// TIA Portal project "FORMING_1500_PLC" (V15) (continued)

REGION Network 7: Q124.4 ON SELAMA 6 DETIK SETELAH I 7.5 ON
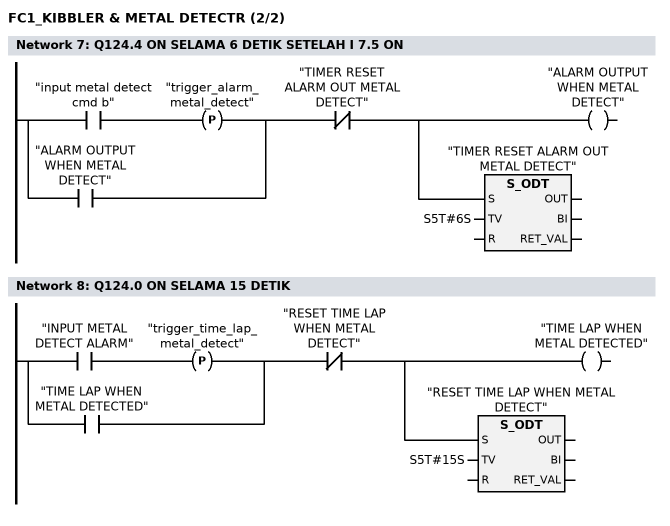
   RUNG wire#powerrail
      Contact( "input metal detect cmd b" )
      P_Trig( "trigger_alarm_metal_detect" )
      wire#w1
      I_Contact( "TIMER RESET ALARM OUT METAL DETECT" )
      wire#w2
      Coil( "ALARM OUTPUT WHEN METAL DETECT" )
   END_RUNG
   RUNG wire#powerrail
      Contact( "ALARM OUTPUT WHEN METAL DETECT" )
   END_RUNG wire#w1
   RUNG wire#w2
      S_ODT(T_NO := "TIMER RESET ALARM OUT METAL DETECT", TV := S5T#6S, R :=, BI =>, RET_VAL =>)
   END_RUNG
   // the same network as SCL:
   #_w1 := "input metal detect cmd b" AND NOT "trigger_alarm_metal_detect";   // rising edge
   "trigger_alarm_metal_detect" := "input metal detect cmd b";
   "ALARM OUTPUT WHEN METAL DETECT" := (#_w1 OR "ALARM OUTPUT WHEN METAL DETECT") AND NOT "TIMER RESET ALARM OUT METAL DETECT";
   #_s5time1 := S_ODT(T_NO := "TIMER RESET ALARM OUT METAL DETECT",
                      S := "ALARM OUTPUT WHEN METAL DETECT",
                      TV := S5T#6S);
END_REGION

REGION Network 8: Q124.0 ON SELAMA 15 DETIK
   RUNG wire#powerrail
      Contact( "INPUT METAL DETECT ALARM" )
      P_Trig( "trigger_time_lap_metal_detect" )
      wire#w1
      I_Contact( "RESET TIME LAP WHEN METAL DETECT" )
      wire#w2
      Coil( "TIME LAP WHEN METAL DETECTED" )
   END_RUNG
   RUNG wire#powerrail
      Contact( "TIME LAP WHEN METAL DETECTED" )
   END_RUNG wire#w1
   RUNG wire#w2
      S_ODT(T_NO := "RESET TIME LAP WHEN METAL DETECT", TV := S5T#15S, R :=, BI =>, RET_VAL =>)
   END_RUNG
   // the same network as SCL:
   #_w1 := "INPUT METAL DETECT ALARM" AND NOT "trigger_time_lap_metal_detect";   // rising edge
   "trigger_time_lap_metal_detect" := "INPUT METAL DETECT ALARM";
   "TIME LAP WHEN METAL DETECTED" := (#_w1 OR "TIME LAP WHEN METAL DETECTED") AND NOT "RESET TIME LAP WHEN METAL DETECT";
   #_s5time1 := S_ODT(T_NO := "RESET TIME LAP WHEN METAL DETECT",
                      S := "TIME LAP WHEN METAL DETECTED",
                      TV := S5T#15S);
END_REGION
END_FUNCTION

FUNCTION "FC2" : Void   // FC2, LAD
{ S7_Optimized_Access := 'FALSE' }
VERSION : 0.1
BEGIN
END_FUNCTION

FUNCTION "FC3_SPEED REFF/ MRV" : Void   // FC3, LAD
TITLE = Speed Refference to inverter
{ S7_Optimized_Access := 'FALSE' }
VERSION : 0.1
BEGIN

REGION Network 1: MAIN REFERENCE VALUE / SPEED REFFERENCE ADDRESS 2
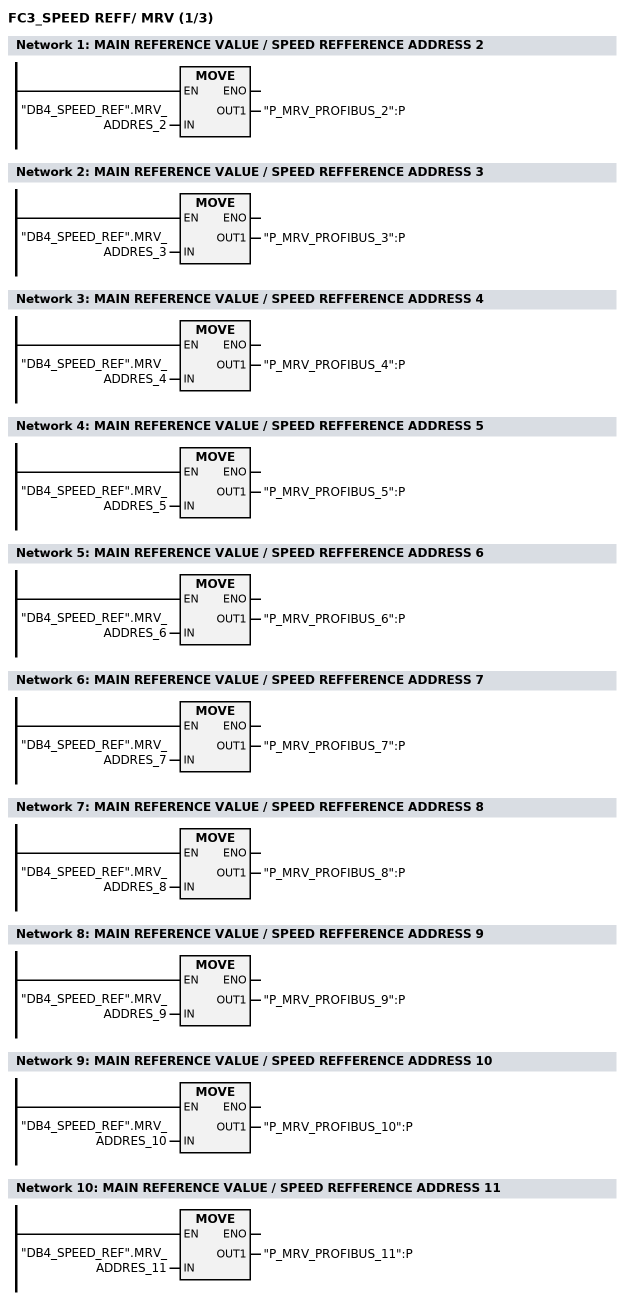
   RUNG wire#powerrail
      { S7_GenerateENO := "TRUE" } Move(in := "DB4_SPEED_REF".MRV_ADDRES_2, out1 => "P_MRV_PROFIBUS_2":P)
   END_RUNG
   // the same network as SCL:
   "P_MRV_PROFIBUS_2":P := "DB4_SPEED_REF".MRV_ADDRES_2;
END_REGION

REGION Network 2: MAIN REFERENCE VALUE / SPEED REFFERENCE ADDRESS 3
   RUNG wire#powerrail
      { S7_GenerateENO := "TRUE" } Move(in := "DB4_SPEED_REF".MRV_ADDRES_3, out1 => "P_MRV_PROFIBUS_3":P)
   END_RUNG
   // the same network as SCL:
   "P_MRV_PROFIBUS_3":P := "DB4_SPEED_REF".MRV_ADDRES_3;
END_REGION

REGION Network 3: MAIN REFERENCE VALUE / SPEED REFFERENCE ADDRESS 4
   RUNG wire#powerrail
      { S7_GenerateENO := "TRUE" } Move(in := "DB4_SPEED_REF".MRV_ADDRES_4, out1 => "P_MRV_PROFIBUS_4":P)
   END_RUNG
   // the same network as SCL:
   "P_MRV_PROFIBUS_4":P := "DB4_SPEED_REF".MRV_ADDRES_4;
END_REGION

REGION Network 4: MAIN REFERENCE VALUE / SPEED REFFERENCE ADDRESS 5
   RUNG wire#powerrail
      { S7_GenerateENO := "TRUE" } Move(in := "DB4_SPEED_REF".MRV_ADDRES_5, out1 => "P_MRV_PROFIBUS_5":P)
   END_RUNG
   // the same network as SCL:
   "P_MRV_PROFIBUS_5":P := "DB4_SPEED_REF".MRV_ADDRES_5;
END_REGION

REGION Network 5: MAIN REFERENCE VALUE / SPEED REFFERENCE ADDRESS 6
   RUNG wire#powerrail
      { S7_GenerateENO := "TRUE" } Move(in := "DB4_SPEED_REF".MRV_ADDRES_6, out1 => "P_MRV_PROFIBUS_6":P)
   END_RUNG
   // the same network as SCL:
   "P_MRV_PROFIBUS_6":P := "DB4_SPEED_REF".MRV_ADDRES_6;
END_REGION

REGION Network 6: MAIN REFERENCE VALUE / SPEED REFFERENCE ADDRESS 7
   RUNG wire#powerrail
      { S7_GenerateENO := "TRUE" } Move(in := "DB4_SPEED_REF".MRV_ADDRES_7, out1 => "P_MRV_PROFIBUS_7":P)
   END_RUNG
   // the same network as SCL:
   "P_MRV_PROFIBUS_7":P := "DB4_SPEED_REF".MRV_ADDRES_7;
END_REGION

REGION Network 7: MAIN REFERENCE VALUE / SPEED REFFERENCE ADDRESS 8
   RUNG wire#powerrail
      { S7_GenerateENO := "TRUE" } Move(in := "DB4_SPEED_REF".MRV_ADDRES_8, out1 => "P_MRV_PROFIBUS_8":P)
   END_RUNG
   // the same network as SCL:
   "P_MRV_PROFIBUS_8":P := "DB4_SPEED_REF".MRV_ADDRES_8;
END_REGION

REGION Network 8: MAIN REFERENCE VALUE / SPEED REFFERENCE ADDRESS 9
   RUNG wire#powerrail
      { S7_GenerateENO := "TRUE" } Move(in := "DB4_SPEED_REF".MRV_ADDRES_9, out1 => "P_MRV_PROFIBUS_9":P)
   END_RUNG
   // the same network as SCL:
   "P_MRV_PROFIBUS_9":P := "DB4_SPEED_REF".MRV_ADDRES_9;
END_REGION

REGION Network 9: MAIN REFERENCE VALUE / SPEED REFFERENCE ADDRESS 10
   RUNG wire#powerrail
      { S7_GenerateENO := "TRUE" } Move(in := "DB4_SPEED_REF".MRV_ADDRES_10, out1 => "P_MRV_PROFIBUS_10":P)
   END_RUNG
   // the same network as SCL:
   "P_MRV_PROFIBUS_10":P := "DB4_SPEED_REF".MRV_ADDRES_10;
END_REGION

REGION Network 10: MAIN REFERENCE VALUE / SPEED REFFERENCE ADDRESS 11
   RUNG wire#powerrail
      { S7_GenerateENO := "TRUE" } Move(in := "DB4_SPEED_REF".MRV_ADDRES_11, out1 => "P_MRV_PROFIBUS_11":P)
   END_RUNG
   // the same network as SCL:
   "P_MRV_PROFIBUS_11":P := "DB4_SPEED_REF".MRV_ADDRES_11;
END_REGION

REGION Network 11: MAIN REFERENCE VALUE / SPEED REFFERENCE ADDRESS 12
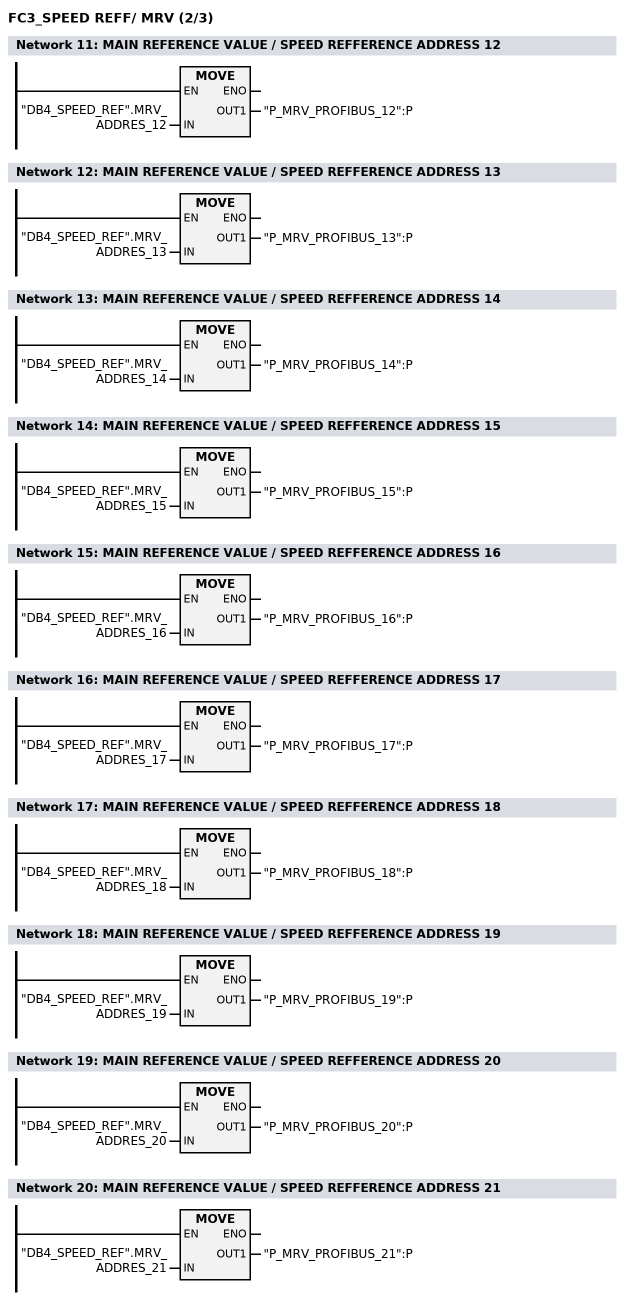
   RUNG wire#powerrail
      { S7_GenerateENO := "TRUE" } Move(in := "DB4_SPEED_REF".MRV_ADDRES_12, out1 => "P_MRV_PROFIBUS_12":P)
   END_RUNG
   // the same network as SCL:
   "P_MRV_PROFIBUS_12":P := "DB4_SPEED_REF".MRV_ADDRES_12;
END_REGION

REGION Network 12: MAIN REFERENCE VALUE / SPEED REFFERENCE ADDRESS 13
   RUNG wire#powerrail
      { S7_GenerateENO := "TRUE" } Move(in := "DB4_SPEED_REF".MRV_ADDRES_13, out1 => "P_MRV_PROFIBUS_13":P)
   END_RUNG
   // the same network as SCL:
   "P_MRV_PROFIBUS_13":P := "DB4_SPEED_REF".MRV_ADDRES_13;
END_REGION

REGION Network 13: MAIN REFERENCE VALUE / SPEED REFFERENCE ADDRESS 14
   RUNG wire#powerrail
      { S7_GenerateENO := "TRUE" } Move(in := "DB4_SPEED_REF".MRV_ADDRES_14, out1 => "P_MRV_PROFIBUS_14":P)
   END_RUNG
   // the same network as SCL:
   "P_MRV_PROFIBUS_14":P := "DB4_SPEED_REF".MRV_ADDRES_14;
END_REGION

REGION Network 14: MAIN REFERENCE VALUE / SPEED REFFERENCE ADDRESS 15
   RUNG wire#powerrail
      { S7_GenerateENO := "TRUE" } Move(in := "DB4_SPEED_REF".MRV_ADDRES_15, out1 => "P_MRV_PROFIBUS_15":P)
   END_RUNG
   // the same network as SCL:
   "P_MRV_PROFIBUS_15":P := "DB4_SPEED_REF".MRV_ADDRES_15;
END_REGION

REGION Network 15: MAIN REFERENCE VALUE / SPEED REFFERENCE ADDRESS 16
   RUNG wire#powerrail
      { S7_GenerateENO := "TRUE" } Move(in := "DB4_SPEED_REF".MRV_ADDRES_16, out1 => "P_MRV_PROFIBUS_16":P)
   END_RUNG
   // the same network as SCL:
   "P_MRV_PROFIBUS_16":P := "DB4_SPEED_REF".MRV_ADDRES_16;
END_REGION

REGION Network 16: MAIN REFERENCE VALUE / SPEED REFFERENCE ADDRESS 17
   RUNG wire#powerrail
      { S7_GenerateENO := "TRUE" } Move(in := "DB4_SPEED_REF".MRV_ADDRES_17, out1 => "P_MRV_PROFIBUS_17":P)
   END_RUNG
   // the same network as SCL:
   "P_MRV_PROFIBUS_17":P := "DB4_SPEED_REF".MRV_ADDRES_17;
END_REGION

REGION Network 17: MAIN REFERENCE VALUE / SPEED REFFERENCE ADDRESS 18
   RUNG wire#powerrail
      { S7_GenerateENO := "TRUE" } Move(in := "DB4_SPEED_REF".MRV_ADDRES_18, out1 => "P_MRV_PROFIBUS_18":P)
   END_RUNG
   // the same network as SCL:
   "P_MRV_PROFIBUS_18":P := "DB4_SPEED_REF".MRV_ADDRES_18;
END_REGION

REGION Network 18: MAIN REFERENCE VALUE / SPEED REFFERENCE ADDRESS 19
   RUNG wire#powerrail
      { S7_GenerateENO := "TRUE" } Move(in := "DB4_SPEED_REF".MRV_ADDRES_19, out1 => "P_MRV_PROFIBUS_19":P)
   END_RUNG
   // the same network as SCL:
   "P_MRV_PROFIBUS_19":P := "DB4_SPEED_REF".MRV_ADDRES_19;
END_REGION

REGION Network 19: MAIN REFERENCE VALUE / SPEED REFFERENCE ADDRESS 20
   RUNG wire#powerrail
      { S7_GenerateENO := "TRUE" } Move(in := "DB4_SPEED_REF".MRV_ADDRES_20, out1 => "P_MRV_PROFIBUS_20":P)
   END_RUNG
   // the same network as SCL:
   "P_MRV_PROFIBUS_20":P := "DB4_SPEED_REF".MRV_ADDRES_20;
END_REGION

REGION Network 20: MAIN REFERENCE VALUE / SPEED REFFERENCE ADDRESS 21
   RUNG wire#powerrail
      { S7_GenerateENO := "TRUE" } Move(in := "DB4_SPEED_REF".MRV_ADDRES_21, out1 => "P_MRV_PROFIBUS_21":P)
   END_RUNG
   // the same network as SCL:
   "P_MRV_PROFIBUS_21":P := "DB4_SPEED_REF".MRV_ADDRES_21;
END_REGION

REGION Network 21: MAIN REFERENCE VALUE / SPEED REFFERENCE ADDRESS 22
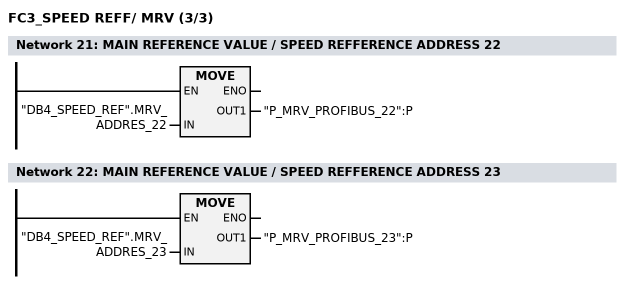
   RUNG wire#powerrail
      { S7_GenerateENO := "TRUE" } Move(in := "DB4_SPEED_REF".MRV_ADDRES_22, out1 => "P_MRV_PROFIBUS_22":P)
   END_RUNG
   // the same network as SCL:
   "P_MRV_PROFIBUS_22":P := "DB4_SPEED_REF".MRV_ADDRES_22;
END_REGION

REGION Network 22: MAIN REFERENCE VALUE / SPEED REFFERENCE ADDRESS 23
   RUNG wire#powerrail
      { S7_GenerateENO := "TRUE" } Move(in := "DB4_SPEED_REF".MRV_ADDRES_23, out1 => "P_MRV_PROFIBUS_23":P)
   END_RUNG
   // the same network as SCL:
   "P_MRV_PROFIBUS_23":P := "DB4_SPEED_REF".MRV_ADDRES_23;
END_REGION
END_FUNCTION

FUNCTION "FC4" : Void   // FC4, LAD
{ S7_Optimized_Access := 'FALSE' }
VERSION : 0.1
BEGIN
END_FUNCTION

FUNCTION "FC5_INC_DEC_A" : Void   // FC5, LAD
TITLE = Increment Decrement inverter 2,13,17,20 & transfer speed from synchron to single
{ S7_Optimized_Access := 'FALSE' }
VERSION : 0.1
   VAR_TEMP   // added for the SCL form of the ladder/FBD networks
      _w1 : Bool;
      _w2 : Bool;
   END_VAR
BEGIN

REGION Network 1: ADDRESS 13 / I 7.0 | Increase Decrease ADDRESS 13
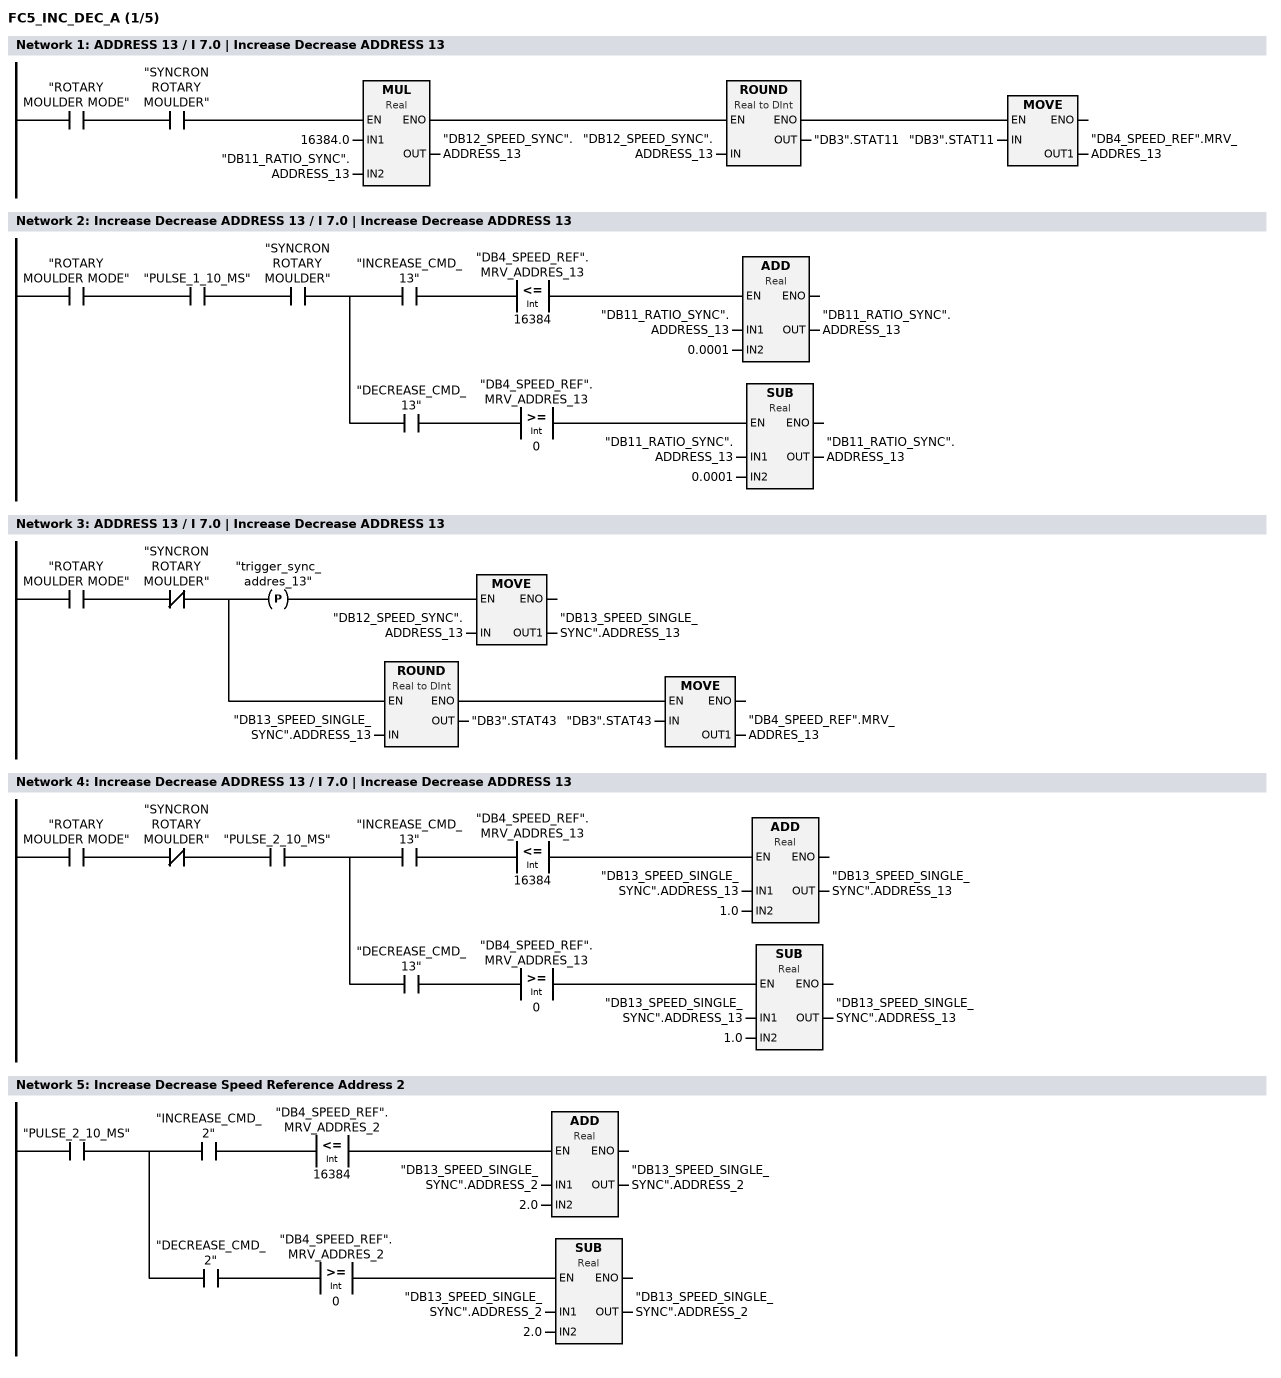
   RUNG wire#powerrail
      Contact( "ROTARY MOULDER MODE" )
      Contact( "SYNCRON ROTARY MOULDER" )
      { S7_Templates := "SrcType := Real"; S7_GenerateENO := "TRUE" } Mul(in1 := 16384.0, in2 := "DB11_RATIO_SYNC".ADDRESS_13, out => "DB12_SPEED_SYNC".ADDRESS_13)
      { S7_Templates := "[SrcType := Real, DestType := DInt]"; S7_GenerateENO := "TRUE" } Round(in := "DB12_SPEED_SYNC".ADDRESS_13, out => "DB3".STAT11)
      { S7_GenerateENO := "TRUE" } Move(in := "DB3".STAT11, out1 => "DB4_SPEED_REF".MRV_ADDRES_13)
   END_RUNG
   // the same network as SCL:
   // ENO of a box is taken as its EN; it also drops when the box reports an error
   IF "ROTARY MOULDER MODE" AND "SYNCRON ROTARY MOULDER" THEN
       "DB12_SPEED_SYNC".ADDRESS_13 := 16384.0 * "DB11_RATIO_SYNC".ADDRESS_13;
       "DB3".STAT11 := ROUND("DB12_SPEED_SYNC".ADDRESS_13);
       "DB4_SPEED_REF".MRV_ADDRES_13 := "DB3".STAT11;
   END_IF;
END_REGION

REGION Network 2: Increase Decrease ADDRESS 13 / I 7.0 | Increase Decrease ADDRESS 13
   RUNG wire#powerrail
      Contact( "ROTARY MOULDER MODE" )
      Contact( "PULSE_1_10_MS" )
      Contact( "SYNCRON ROTARY MOULDER" )
      wire#w1
      Contact( "INCREASE_CMD_13" )
      { S7_Templates := "SrcType := Int" } LE_Contact(in1 := "DB4_SPEED_REF".MRV_ADDRES_13, in2 := 16384)
      { S7_Templates := "SrcType := Real"; S7_GenerateENO := "TRUE" } Add(in1 := "DB11_RATIO_SYNC".ADDRESS_13, in2 := 0.0001, out => "DB11_RATIO_SYNC".ADDRESS_13)
   END_RUNG
   RUNG wire#w1
      Contact( "DECREASE_CMD_13" )
      { S7_Templates := "SrcType := Int" } GE_Contact(in1 := "DB4_SPEED_REF".MRV_ADDRES_13, in2 := 0)
      { S7_Templates := "SrcType := Real"; S7_GenerateENO := "TRUE" } Sub(in1 := "DB11_RATIO_SYNC".ADDRESS_13, in2 := 0.0001, out => "DB11_RATIO_SYNC".ADDRESS_13)
   END_RUNG
   // the same network as SCL:
   #_w1 := "ROTARY MOULDER MODE" AND "PULSE_1_10_MS" AND "SYNCRON ROTARY MOULDER";
   IF #_w1 AND "INCREASE_CMD_13" AND ("DB4_SPEED_REF".MRV_ADDRES_13 <= 16384) THEN
       "DB11_RATIO_SYNC".ADDRESS_13 := "DB11_RATIO_SYNC".ADDRESS_13 + 0.0001;
   END_IF;
   IF #_w1 AND "DECREASE_CMD_13" AND ("DB4_SPEED_REF".MRV_ADDRES_13 >= 0) THEN
       "DB11_RATIO_SYNC".ADDRESS_13 := "DB11_RATIO_SYNC".ADDRESS_13 - 0.0001;
   END_IF;
END_REGION

REGION Network 3: ADDRESS 13 / I 7.0 | Increase Decrease ADDRESS 13
   RUNG wire#powerrail
      Contact( "ROTARY MOULDER MODE" )
      I_Contact( "SYNCRON ROTARY MOULDER" )
      wire#w1
      P_Trig( "trigger_sync_addres_13" )
      { S7_GenerateENO := "TRUE" } Move(in := "DB12_SPEED_SYNC".ADDRESS_13, out1 => "DB13_SPEED_SINGLE_SYNC".ADDRESS_13)
   END_RUNG
   RUNG wire#w1
      { S7_Templates := "[SrcType := Real, DestType := DInt]"; S7_GenerateENO := "TRUE" } Round(in := "DB13_SPEED_SINGLE_SYNC".ADDRESS_13, out => "DB3".STAT43)
      { S7_GenerateENO := "TRUE" } Move(in := "DB3".STAT43, out1 => "DB4_SPEED_REF".MRV_ADDRES_13)
   END_RUNG
   // the same network as SCL:
   // ENO of a box is taken as its EN; it also drops when the box reports an error
   #_w1 := "ROTARY MOULDER MODE" AND NOT "SYNCRON ROTARY MOULDER";
   #_w2 := #_w1 AND NOT "trigger_sync_addres_13";   // rising edge
   "trigger_sync_addres_13" := #_w1;
   IF #_w2 THEN "DB13_SPEED_SINGLE_SYNC".ADDRESS_13 := "DB12_SPEED_SYNC".ADDRESS_13; END_IF;
   IF #_w1 THEN
       "DB3".STAT43 := ROUND("DB13_SPEED_SINGLE_SYNC".ADDRESS_13);
       "DB4_SPEED_REF".MRV_ADDRES_13 := "DB3".STAT43;
   END_IF;
END_REGION

REGION Network 4: Increase Decrease ADDRESS 13 / I 7.0 | Increase Decrease ADDRESS 13
   RUNG wire#powerrail
      Contact( "ROTARY MOULDER MODE" )
      I_Contact( "SYNCRON ROTARY MOULDER" )
      Contact( "PULSE_2_10_MS" )
      wire#w1
      Contact( "INCREASE_CMD_13" )
      { S7_Templates := "SrcType := Int" } LE_Contact(in1 := "DB4_SPEED_REF".MRV_ADDRES_13, in2 := 16384)
      { S7_Templates := "SrcType := Real"; S7_GenerateENO := "TRUE" } Add(in1 := "DB13_SPEED_SINGLE_SYNC".ADDRESS_13, in2 := 1.0, out => "DB13_SPEED_SINGLE_SYNC".ADDRESS_13)
   END_RUNG
   RUNG wire#w1
      Contact( "DECREASE_CMD_13" )
      { S7_Templates := "SrcType := Int" } GE_Contact(in1 := "DB4_SPEED_REF".MRV_ADDRES_13, in2 := 0)
      { S7_Templates := "SrcType := Real"; S7_GenerateENO := "TRUE" } Sub(in1 := "DB13_SPEED_SINGLE_SYNC".ADDRESS_13, in2 := 1.0, out => "DB13_SPEED_SINGLE_SYNC".ADDRESS_13)
   END_RUNG
   // the same network as SCL:
   #_w1 := "ROTARY MOULDER MODE" AND NOT "SYNCRON ROTARY MOULDER" AND "PULSE_2_10_MS";
   IF #_w1 AND "INCREASE_CMD_13" AND ("DB4_SPEED_REF".MRV_ADDRES_13 <= 16384) THEN
       "DB13_SPEED_SINGLE_SYNC".ADDRESS_13 := "DB13_SPEED_SINGLE_SYNC".ADDRESS_13 + 1.0;
   END_IF;
   IF #_w1 AND "DECREASE_CMD_13" AND ("DB4_SPEED_REF".MRV_ADDRES_13 >= 0) THEN
       "DB13_SPEED_SINGLE_SYNC".ADDRESS_13 := "DB13_SPEED_SINGLE_SYNC".ADDRESS_13 - 1.0;
   END_IF;
END_REGION

REGION Network 5: Increase Decrease Speed Reference Address 2
   RUNG wire#powerrail
      Contact( "PULSE_2_10_MS" )
      wire#w1
      Contact( "INCREASE_CMD_2" )
      { S7_Templates := "SrcType := Int" } LE_Contact(in1 := "DB4_SPEED_REF".MRV_ADDRES_2, in2 := 16384)
      { S7_Templates := "SrcType := Real"; S7_GenerateENO := "TRUE" } Add(in1 := "DB13_SPEED_SINGLE_SYNC".ADDRESS_2, in2 := 2.0, out => "DB13_SPEED_SINGLE_SYNC".ADDRESS_2)
   END_RUNG
   RUNG wire#w1
      Contact( "DECREASE_CMD_2" )
      { S7_Templates := "SrcType := Int" } GE_Contact(in1 := "DB4_SPEED_REF".MRV_ADDRES_2, in2 := 0)
      { S7_Templates := "SrcType := Real"; S7_GenerateENO := "TRUE" } Sub(in1 := "DB13_SPEED_SINGLE_SYNC".ADDRESS_2, in2 := 2.0, out => "DB13_SPEED_SINGLE_SYNC".ADDRESS_2)
   END_RUNG
   // the same network as SCL:
   IF "PULSE_2_10_MS" AND "INCREASE_CMD_2" AND ("DB4_SPEED_REF".MRV_ADDRES_2 <= 16384) THEN
       "DB13_SPEED_SINGLE_SYNC".ADDRESS_2 := "DB13_SPEED_SINGLE_SYNC".ADDRESS_2 + 2.0;
   END_IF;
   IF "PULSE_2_10_MS" AND "DECREASE_CMD_2" AND ("DB4_SPEED_REF".MRV_ADDRES_2 >= 0) THEN
       "DB13_SPEED_SINGLE_SYNC".ADDRESS_2 := "DB13_SPEED_SINGLE_SYNC".ADDRESS_2 - 2.0;
   END_IF;
END_REGION

REGION Network 6: Control Speed Address 2 / Increase Decrease Speed Reference Address 2
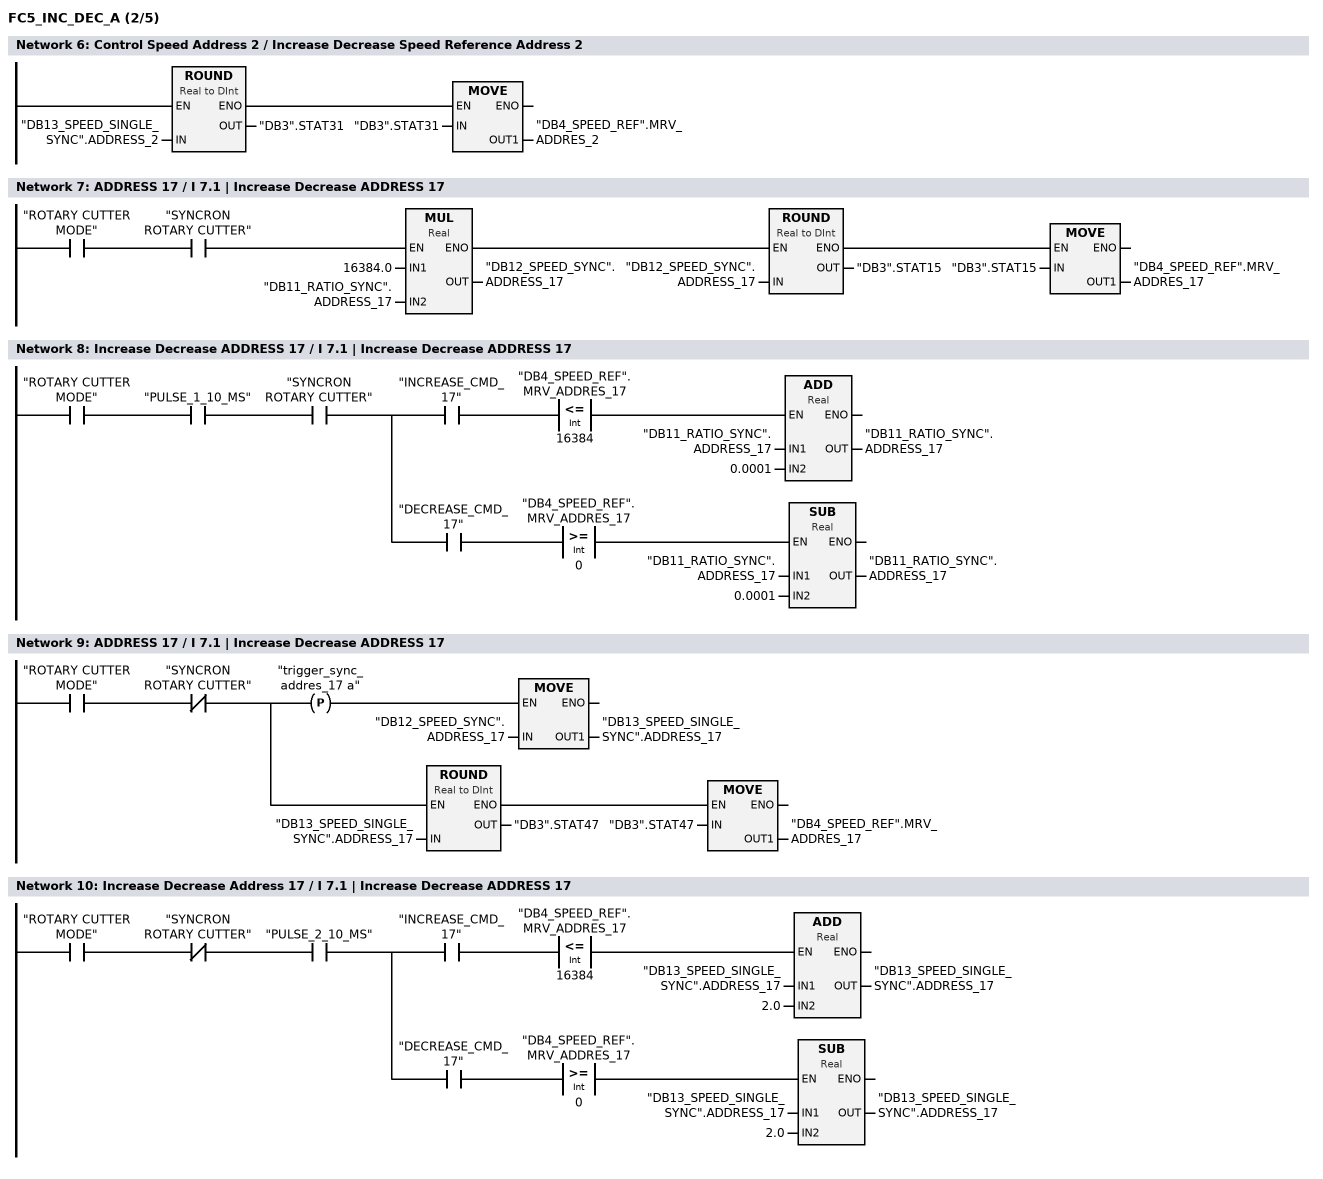
   RUNG wire#powerrail
      { S7_Templates := "[SrcType := Real, DestType := DInt]"; S7_GenerateENO := "TRUE" } Round(in := "DB13_SPEED_SINGLE_SYNC".ADDRESS_2, out => "DB3".STAT31)
      { S7_GenerateENO := "TRUE" } Move(in := "DB3".STAT31, out1 => "DB4_SPEED_REF".MRV_ADDRES_2)
   END_RUNG
   // the same network as SCL:
   // ENO of a box is taken as its EN; it also drops when the box reports an error
   "DB3".STAT31 := ROUND("DB13_SPEED_SINGLE_SYNC".ADDRESS_2);
   "DB4_SPEED_REF".MRV_ADDRES_2 := "DB3".STAT31;
END_REGION

REGION Network 7: ADDRESS 17 / I 7.1 | Increase Decrease ADDRESS 17
   RUNG wire#powerrail
      Contact( "ROTARY CUTTER MODE" )
      Contact( "SYNCRON ROTARY CUTTER" )
      { S7_Templates := "SrcType := Real"; S7_GenerateENO := "TRUE" } Mul(in1 := 16384.0, in2 := "DB11_RATIO_SYNC".ADDRESS_17, out => "DB12_SPEED_SYNC".ADDRESS_17)
      { S7_Templates := "[SrcType := Real, DestType := DInt]"; S7_GenerateENO := "TRUE" } Round(in := "DB12_SPEED_SYNC".ADDRESS_17, out => "DB3".STAT15)
      { S7_GenerateENO := "TRUE" } Move(in := "DB3".STAT15, out1 => "DB4_SPEED_REF".MRV_ADDRES_17)
   END_RUNG
   // the same network as SCL:
   // ENO of a box is taken as its EN; it also drops when the box reports an error
   IF "ROTARY CUTTER MODE" AND "SYNCRON ROTARY CUTTER" THEN
       "DB12_SPEED_SYNC".ADDRESS_17 := 16384.0 * "DB11_RATIO_SYNC".ADDRESS_17;
       "DB3".STAT15 := ROUND("DB12_SPEED_SYNC".ADDRESS_17);
       "DB4_SPEED_REF".MRV_ADDRES_17 := "DB3".STAT15;
   END_IF;
END_REGION

REGION Network 8: Increase Decrease ADDRESS 17 / I 7.1 | Increase Decrease ADDRESS 17
   RUNG wire#powerrail
      Contact( "ROTARY CUTTER MODE" )
      Contact( "PULSE_1_10_MS" )
      Contact( "SYNCRON ROTARY CUTTER" )
      wire#w1
      Contact( "INCREASE_CMD_17" )
      { S7_Templates := "SrcType := Int" } LE_Contact(in1 := "DB4_SPEED_REF".MRV_ADDRES_17, in2 := 16384)
      { S7_Templates := "SrcType := Real"; S7_GenerateENO := "TRUE" } Add(in1 := "DB11_RATIO_SYNC".ADDRESS_17, in2 := 0.0001, out => "DB11_RATIO_SYNC".ADDRESS_17)
   END_RUNG
   RUNG wire#w1
      Contact( "DECREASE_CMD_17" )
      { S7_Templates := "SrcType := Int" } GE_Contact(in1 := "DB4_SPEED_REF".MRV_ADDRES_17, in2 := 0)
      { S7_Templates := "SrcType := Real"; S7_GenerateENO := "TRUE" } Sub(in1 := "DB11_RATIO_SYNC".ADDRESS_17, in2 := 0.0001, out => "DB11_RATIO_SYNC".ADDRESS_17)
   END_RUNG
   // the same network as SCL:
   #_w1 := "ROTARY CUTTER MODE" AND "PULSE_1_10_MS" AND "SYNCRON ROTARY CUTTER";
   IF #_w1 AND "INCREASE_CMD_17" AND ("DB4_SPEED_REF".MRV_ADDRES_17 <= 16384) THEN
       "DB11_RATIO_SYNC".ADDRESS_17 := "DB11_RATIO_SYNC".ADDRESS_17 + 0.0001;
   END_IF;
   IF #_w1 AND "DECREASE_CMD_17" AND ("DB4_SPEED_REF".MRV_ADDRES_17 >= 0) THEN
       "DB11_RATIO_SYNC".ADDRESS_17 := "DB11_RATIO_SYNC".ADDRESS_17 - 0.0001;
   END_IF;
END_REGION

REGION Network 9: ADDRESS 17 / I 7.1 | Increase Decrease ADDRESS 17
   RUNG wire#powerrail
      Contact( "ROTARY CUTTER MODE" )
      I_Contact( "SYNCRON ROTARY CUTTER" )
      wire#w1
      P_Trig( "trigger_sync_addres_17 a" )
      { S7_GenerateENO := "TRUE" } Move(in := "DB12_SPEED_SYNC".ADDRESS_17, out1 => "DB13_SPEED_SINGLE_SYNC".ADDRESS_17)
   END_RUNG
   RUNG wire#w1
      { S7_Templates := "[SrcType := Real, DestType := DInt]"; S7_GenerateENO := "TRUE" } Round(in := "DB13_SPEED_SINGLE_SYNC".ADDRESS_17, out => "DB3".STAT47)
      { S7_GenerateENO := "TRUE" } Move(in := "DB3".STAT47, out1 => "DB4_SPEED_REF".MRV_ADDRES_17)
   END_RUNG
   // the same network as SCL:
   // ENO of a box is taken as its EN; it also drops when the box reports an error
   #_w1 := "ROTARY CUTTER MODE" AND NOT "SYNCRON ROTARY CUTTER";
   #_w2 := #_w1 AND NOT "trigger_sync_addres_17 a";   // rising edge
   "trigger_sync_addres_17 a" := #_w1;
   IF #_w2 THEN "DB13_SPEED_SINGLE_SYNC".ADDRESS_17 := "DB12_SPEED_SYNC".ADDRESS_17; END_IF;
   IF #_w1 THEN
       "DB3".STAT47 := ROUND("DB13_SPEED_SINGLE_SYNC".ADDRESS_17);
       "DB4_SPEED_REF".MRV_ADDRES_17 := "DB3".STAT47;
   END_IF;
END_REGION

REGION Network 10: Increase Decrease Address 17 / I 7.1 | Increase Decrease ADDRESS 17
   RUNG wire#powerrail
      Contact( "ROTARY CUTTER MODE" )
      I_Contact( "SYNCRON ROTARY CUTTER" )
      Contact( "PULSE_2_10_MS" )
      wire#w1
      Contact( "INCREASE_CMD_17" )
      { S7_Templates := "SrcType := Int" } LE_Contact(in1 := "DB4_SPEED_REF".MRV_ADDRES_17, in2 := 16384)
      { S7_Templates := "SrcType := Real"; S7_GenerateENO := "TRUE" } Add(in1 := "DB13_SPEED_SINGLE_SYNC".ADDRESS_17, in2 := 2.0, out => "DB13_SPEED_SINGLE_SYNC".ADDRESS_17)
   END_RUNG
   RUNG wire#w1
      Contact( "DECREASE_CMD_17" )
      { S7_Templates := "SrcType := Int" } GE_Contact(in1 := "DB4_SPEED_REF".MRV_ADDRES_17, in2 := 0)
      { S7_Templates := "SrcType := Real"; S7_GenerateENO := "TRUE" } Sub(in1 := "DB13_SPEED_SINGLE_SYNC".ADDRESS_17, in2 := 2.0, out => "DB13_SPEED_SINGLE_SYNC".ADDRESS_17)
   END_RUNG
   // the same network as SCL:
   #_w1 := "ROTARY CUTTER MODE" AND NOT "SYNCRON ROTARY CUTTER" AND "PULSE_2_10_MS";
   IF #_w1 AND "INCREASE_CMD_17" AND ("DB4_SPEED_REF".MRV_ADDRES_17 <= 16384) THEN
       "DB13_SPEED_SINGLE_SYNC".ADDRESS_17 := "DB13_SPEED_SINGLE_SYNC".ADDRESS_17 + 2.0;
   END_IF;
   IF #_w1 AND "DECREASE_CMD_17" AND ("DB4_SPEED_REF".MRV_ADDRES_17 >= 0) THEN
       "DB13_SPEED_SINGLE_SYNC".ADDRESS_17 := "DB13_SPEED_SINGLE_SYNC".ADDRESS_17 - 2.0;
   END_IF;
END_REGION

REGION Network 11: Increase Decrease Address 20 / I 7.0 / I 7.1 |Increase Decrease Address 20